// TIA Portal project "ESTHER_Gas_v4.0_4" (V13) (continued)
       #DATA_ADDR := "MB_AD_COUNTER_RST_ENABL";
       #DATA_INT_PTR.DATA[0] := "MB_VAL_COUNT_RST_ENABL";
   END_IF;
   IF #"STEP" = 44 THEN
       #DATA_ADDR := "MB_AD_COUNTER_UNIT_IDX";
       #DATA_INT_PTR.DATA[0] := 0;   // Unit: ln
   END_IF;
   IF #"STEP" = 45 THEN
       #DATA_ADDR := "MB_AD_COUNTER_SP_MODE";
       #DATA_INT_PTR.DATA[0] := "MB_VAL_COUNT_SP_MODE_CHANGE";
   END_IF;
   IF #"STEP" = 46 THEN
       #DATA_ADDR := "MB_AD_COUNTER_NEW_SP";
       #DATA_INT_PTR.DATA[0] := 0;
   END_IF;
   IF #"STEP" = 47 THEN
       #DATA_ADDR := "MB_AD_RESET";
       #DATA_INT_PTR.DATA[0] := 0;
   END_IF;
   IF #"STEP" = 48 THEN
       #DATA_ADDR := "MB_AD_RESET";
       #DATA_INT_PTR.DATA[0] := 3;
   END_IF;
   IF #"STEP" = 49 THEN
       #DATA_ADDR := "MB_AD_COUNTER_MODE";
       #DATA_INT_PTR.DATA[0] := "MB_VAL_COUNT_MODE_UP_LIMIT";
   END_IF;
   IF #"STEP" = 50 THEN
       #MB_MODE := 1;
       #DATA_LEN := 1;
       #DATA_ADDR := #MB_AD_CONTROL_MODE;
       #DATA_INT_PTR.DATA[0] := #MFC_MODE_SP;   // SET ControlMode
   END_IF;
   IF #"STEP" = 60 THEN
       #MB_MODE := 1;
       #DATA_LEN := 1;
       #DATA_ADDR := #MB_AD_CONTROL_MODE;
       #DATA_INT_PTR.DATA[0] := 0;   // SET ControlMode Bus
   END_IF;
   IF #"STEP" = 63 THEN
       #MB_MODE := 1;
       #DATA_LEN := 1;
       #DATA_ADDR := #MB_AD_CONTROL_MODE;
       #DATA_INT_PTR.DATA[0] := 3;   // SET ControlMode Close
   END_IF;
   IF #"STEP" = 68 THEN
       #MB_MODE := 1;
       #DATA_LEN := 1;
       #DATA_ADDR := #MB_AD_CONTROL_MODE;
       #DATA_INT_PTR.DATA[0] := 8;   // SET ControlMode Open
   END_IF;
   IF #"STEP" = 80 THEN
       #MB_MODE := 1;
       #DATA_LEN := 1;
       #DATA_ADDR := "MB_AD_SETPOINT";
       #DATA_INT_PTR.DATA[0] := #MFC_Setpoint;   // Set Setpoint
   END_IF;
END_REGION
END_FUNCTION_BLOCK

FUNCTION_BLOCK "ETAPA_1_HE_NOK"   // FB3, LAD
{ S7_Optimized_Access := 'FALSE' }
VERSION : 0.1
// Inertização da Câmara de testes com Helio.
BEGIN

REGION Network 1
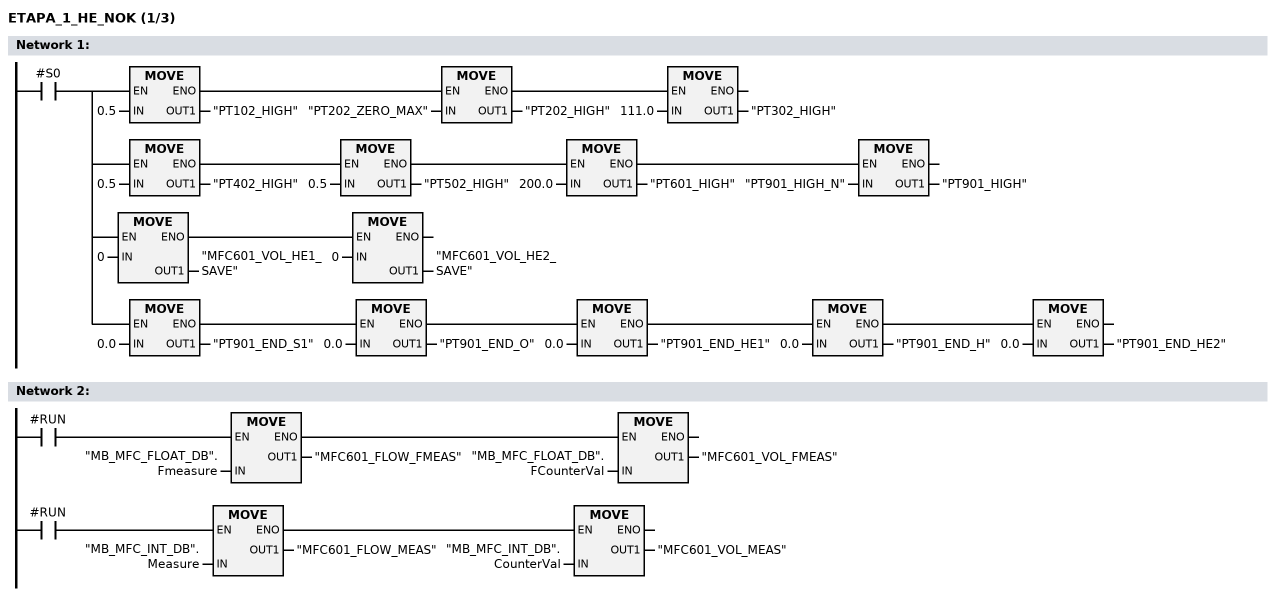
   RUNG wire#powerrail
      Contact( #S0 )
      wire#w1
      { S7_GenerateENO := "TRUE" } Move(in := 0.5, out1 => "PT102_HIGH")
      { S7_GenerateENO := "TRUE" } Move(in := "PT202_ZERO_MAX", out1 => "PT202_HIGH")
      { S7_GenerateENO := "TRUE" } Move(in := 111.0, out1 => "PT302_HIGH")
   END_RUNG
   RUNG wire#w1
      { S7_GenerateENO := "TRUE" } Move(in := 0.5, out1 => "PT402_HIGH")
      { S7_GenerateENO := "TRUE" } Move(in := 0.5, out1 => "PT502_HIGH")
      { S7_GenerateENO := "TRUE" } Move(in := 200.0, out1 => "PT601_HIGH")
      { S7_GenerateENO := "TRUE" } Move(in := "PT901_HIGH_N", out1 => "PT901_HIGH")
   END_RUNG
   RUNG wire#w1
      { S7_GenerateENO := "TRUE" } Move(in := 0, out1 => "MFC601_VOL_HE1_SAVE")
      { S7_GenerateENO := "TRUE" } Move(in := 0, out1 => "MFC601_VOL_HE2_SAVE")
   END_RUNG
   RUNG wire#w1
      { S7_GenerateENO := "TRUE" } Move(in := 0.0, out1 => "PT901_END_S1")
      { S7_GenerateENO := "TRUE" } Move(in := 0.0, out1 => "PT901_END_O")
      { S7_GenerateENO := "TRUE" } Move(in := 0.0, out1 => "PT901_END_HE1")
      { S7_GenerateENO := "TRUE" } Move(in := 0.0, out1 => "PT901_END_H")
      { S7_GenerateENO := "TRUE" } Move(in := 0.0, out1 => "PT901_END_HE2")
   END_RUNG
   // the same network as SCL:
   // ENO of a box is taken as its EN; it also drops when the box reports an error
   IF #S0 THEN
       "PT102_HIGH" := 0.5;
       "PT202_HIGH" := "PT202_ZERO_MAX";
       "PT302_HIGH" := 111.0;
       "PT402_HIGH" := 0.5;
       "PT502_HIGH" := 0.5;
       "PT601_HIGH" := 200.0;
       "PT901_HIGH" := "PT901_HIGH_N";
       "MFC601_VOL_HE1_SAVE" := 0;
       "MFC601_VOL_HE2_SAVE" := 0;
       "PT901_END_S1" := 0.0;
       "PT901_END_O" := 0.0;
       "PT901_END_HE1" := 0.0;
       "PT901_END_H" := 0.0;
       "PT901_END_HE2" := 0.0;
   END_IF;
END_REGION

REGION Network 2
   RUNG wire#powerrail
      Contact( #RUN )
      { S7_GenerateENO := "TRUE" } Move(in := "MB_MFC_FLOAT_DB".Fmeasure, out1 => "MFC601_FLOW_FMEAS")
      { S7_GenerateENO := "TRUE" } Move(in := "MB_MFC_FLOAT_DB".FCounterVal, out1 => "MFC601_VOL_FMEAS")
   END_RUNG
   RUNG wire#powerrail
      Contact( #RUN )
      { S7_GenerateENO := "TRUE" } Move(in := "MB_MFC_INT_DB".Measure, out1 => "MFC601_FLOW_MEAS")
      { S7_GenerateENO := "TRUE" } Move(in := "MB_MFC_INT_DB".CounterVal, out1 => "MFC601_VOL_MEAS")
   END_RUNG
   // the same network as SCL:
   // ENO of a box is taken as its EN; it also drops when the box reports an error
   IF #RUN THEN
       "MFC601_FLOW_FMEAS" := "MB_MFC_FLOAT_DB".Fmeasure;
       "MFC601_VOL_FMEAS" := "MB_MFC_FLOAT_DB".FCounterVal;
       "MFC601_FLOW_MEAS" := "MB_MFC_INT_DB".Measure;
       "MFC601_VOL_MEAS" := "MB_MFC_INT_DB".CounterVal;
   END_IF;
END_REGION

REGION Network 3
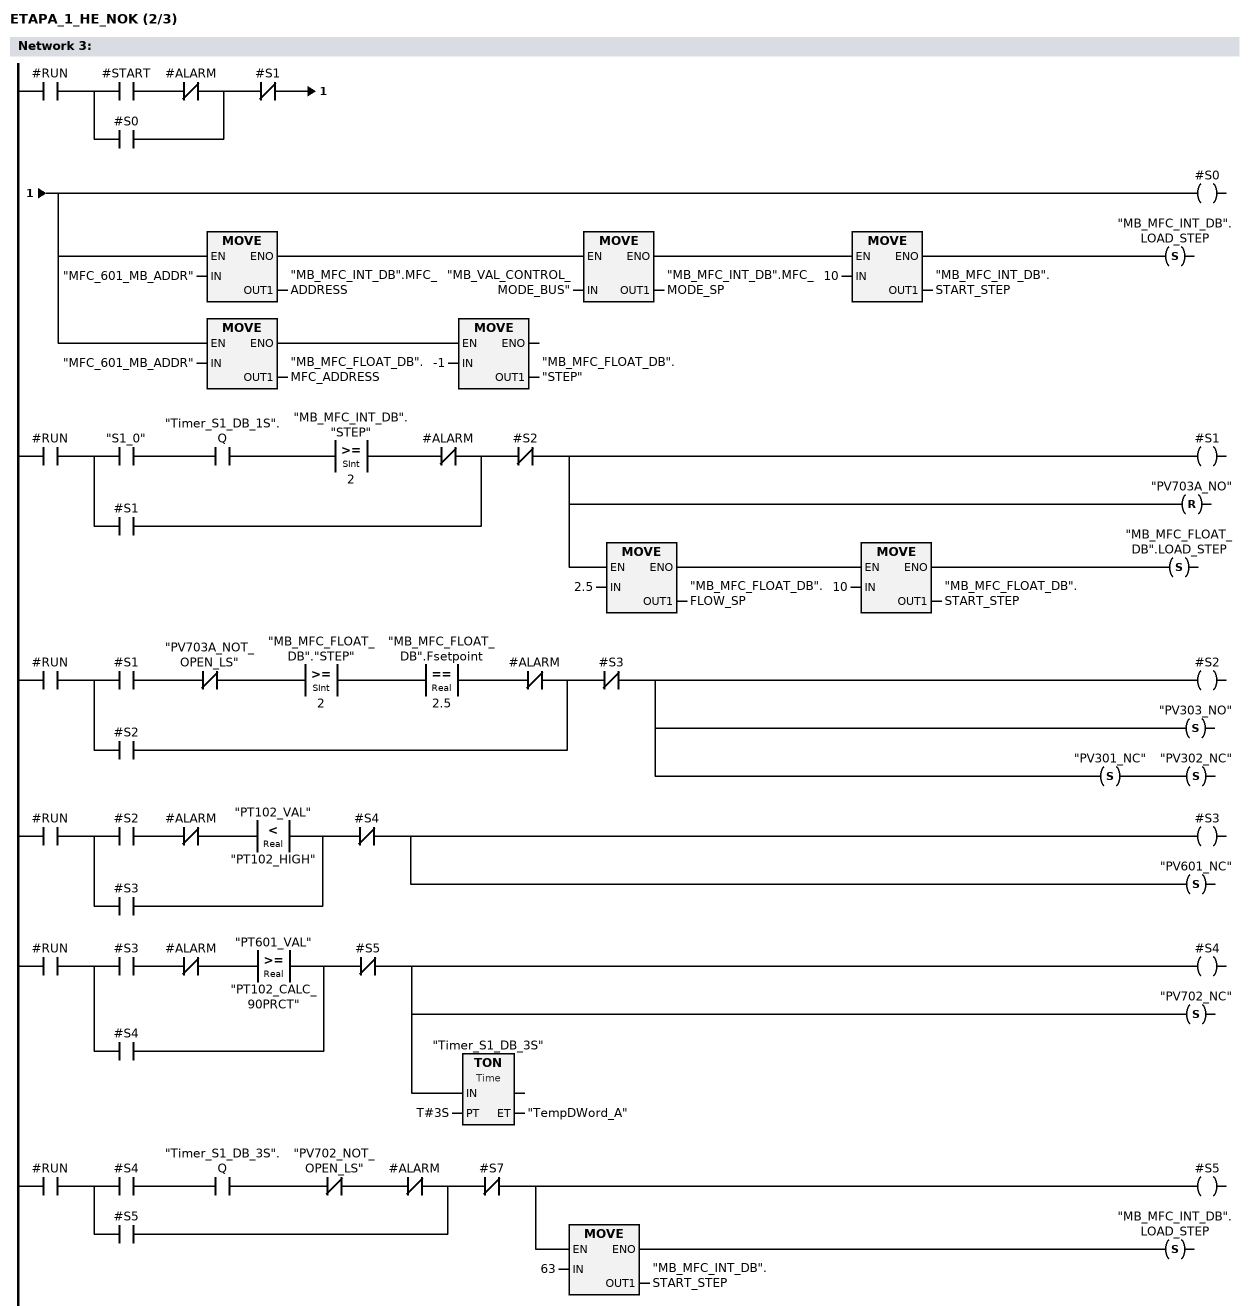
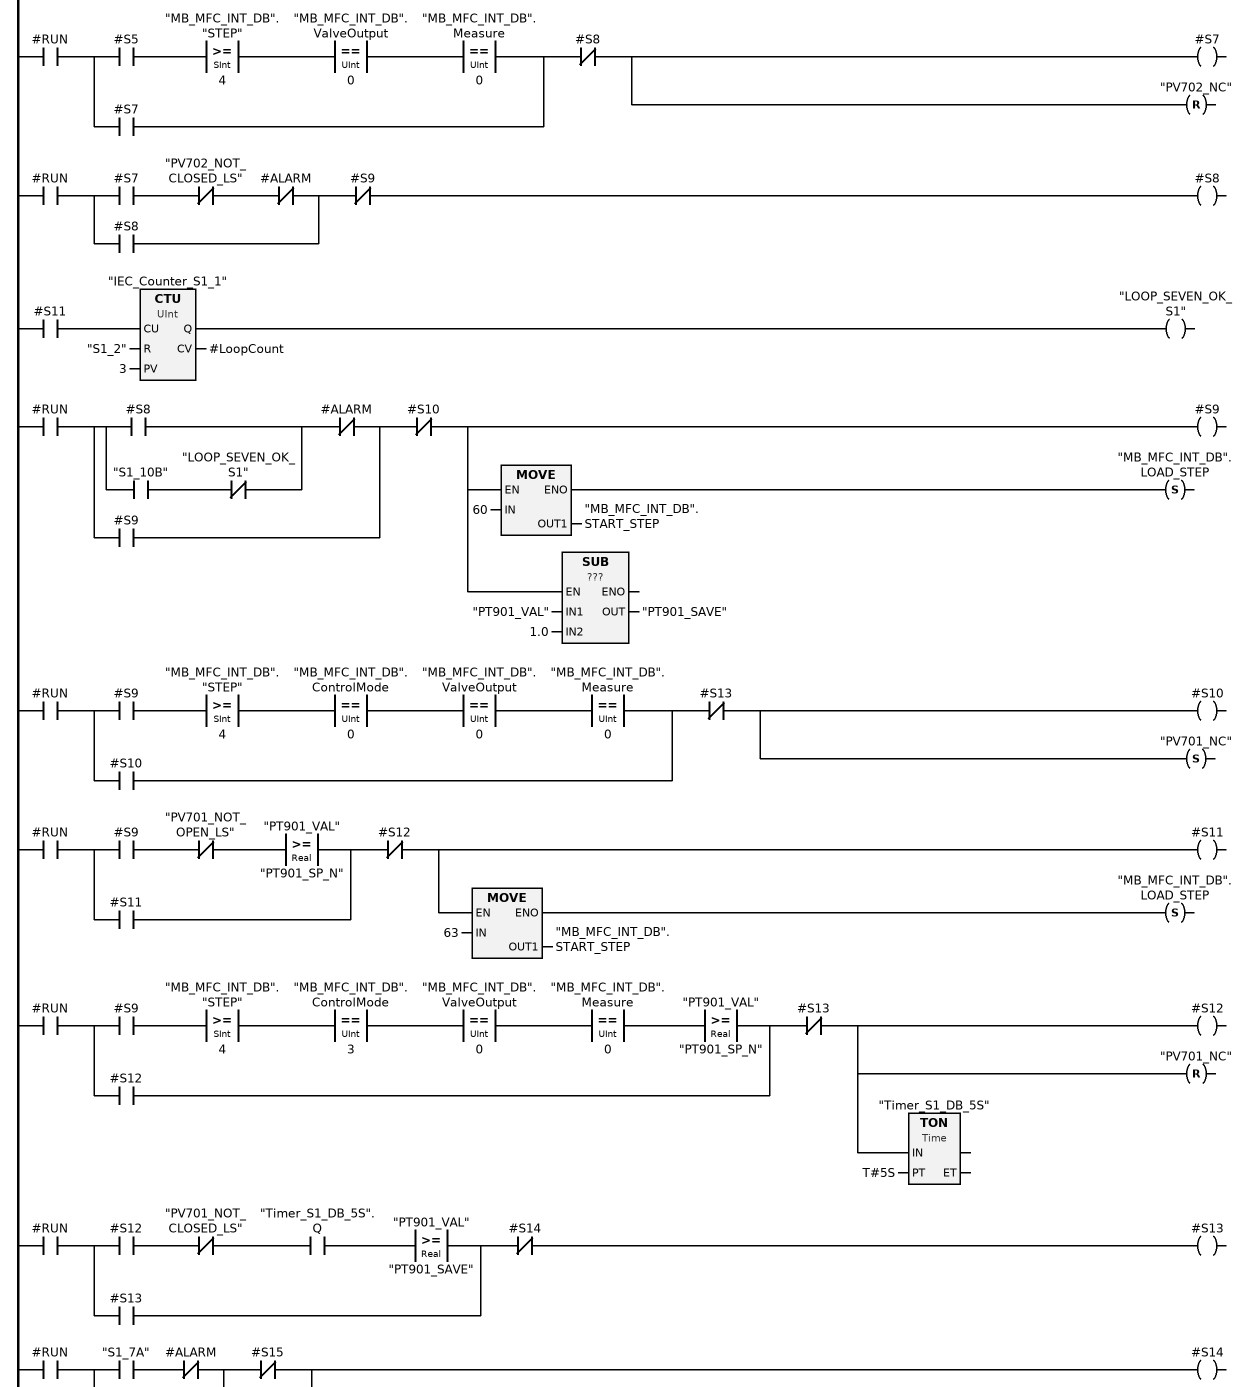
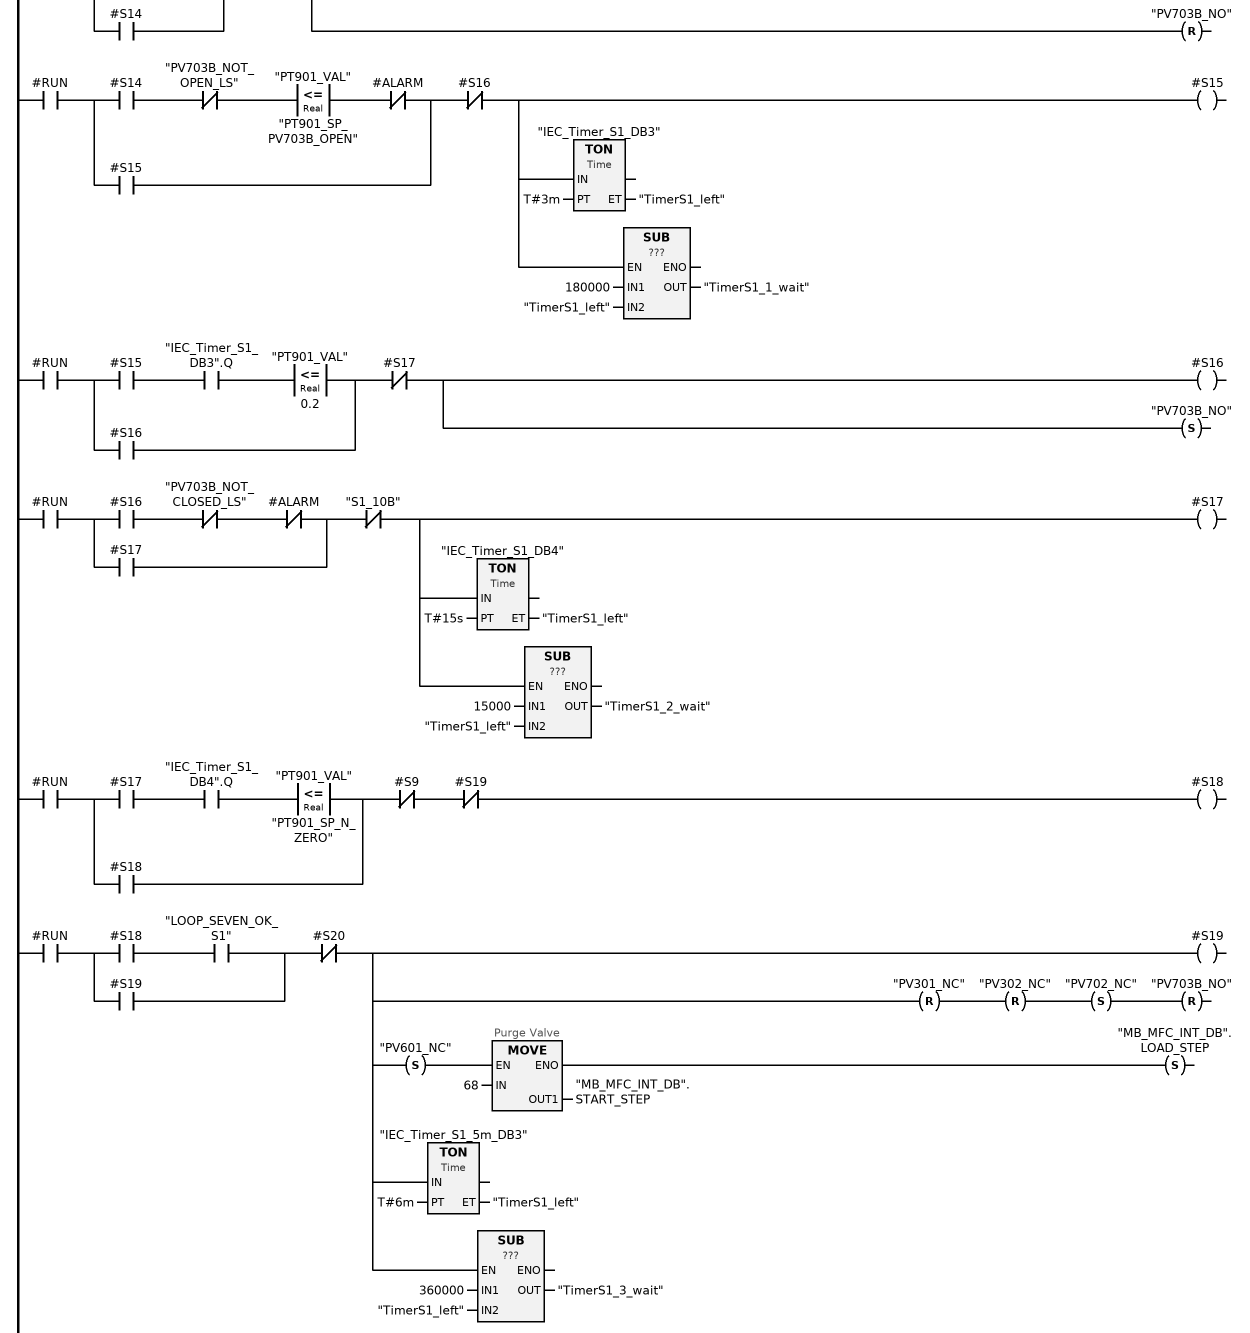
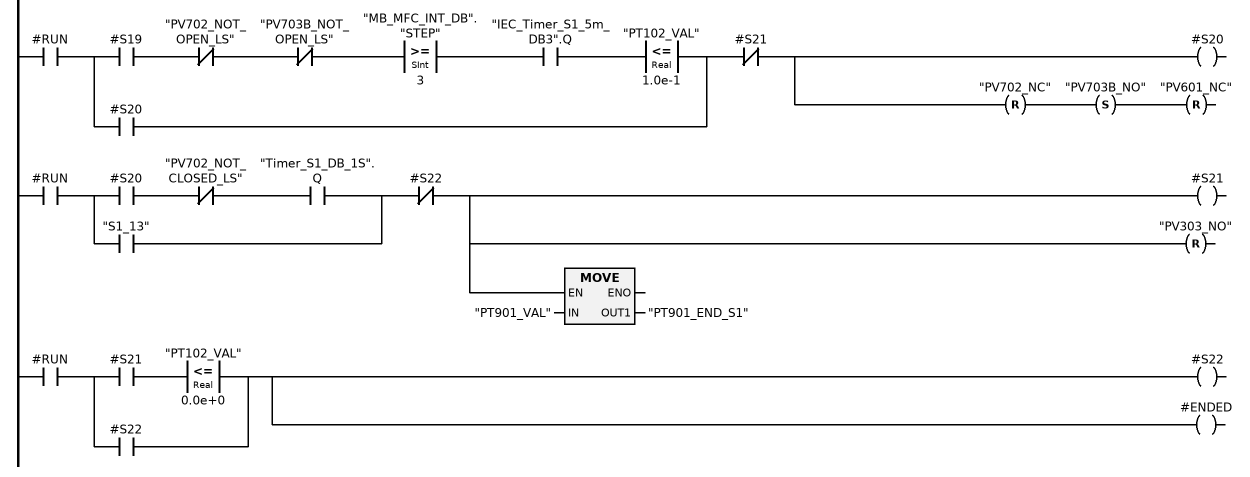
   #S0 := #RUN AND ((#START AND NOT #ALARM) OR #S0) AND NOT #S1;
   IF #S0 THEN
       "MB_MFC_INT_DB".MFC_ADDRESS := "MFC_601_MB_ADDR";
       "MB_MFC_INT_DB".MFC_MODE_SP := "MB_VAL_CONTROL_MODE_BUS";
       "MB_MFC_INT_DB".START_STEP := 10;
       "MB_MFC_INT_DB".LOAD_STEP := TRUE;
       "MB_MFC_FLOAT_DB".MFC_ADDRESS := "MFC_601_MB_ADDR";
       "MB_MFC_FLOAT_DB"."STEP" := -1;
   END_IF;
   #S1 := #RUN AND (("S1_0" AND "Timer_S1_DB_1S".Q AND ("MB_MFC_INT_DB"."STEP" >= 2) AND NOT #ALARM) OR #S1) AND NOT #S2;
   IF #S1 THEN
       "PV703A_NO" := FALSE;
       "MB_MFC_FLOAT_DB".FLOW_SP := 2.5;
       "MB_MFC_FLOAT_DB".START_STEP := 10;
       "MB_MFC_FLOAT_DB".LOAD_STEP := TRUE;
   END_IF;
   #S2 := #RUN AND ((#S1 AND NOT "PV703A_NOT_OPEN_LS" AND ("MB_MFC_FLOAT_DB"."STEP" >= 2) AND ("MB_MFC_FLOAT_DB".Fsetpoint = 2.5) AND NOT #ALARM) OR #S2) AND NOT #S3;
   IF #S2 THEN
       "PV303_NO" := TRUE;
       "PV301_NC" := TRUE;
       "PV302_NC" := TRUE;
   END_IF;
   #S3 := #RUN AND ((#S2 AND NOT #ALARM AND ("PT102_VAL" < "PT102_HIGH")) OR #S3) AND NOT #S4;
   IF #S3 THEN "PV601_NC" := TRUE; END_IF;
   #S4 := #RUN AND ((#S3 AND NOT #ALARM AND ("PT601_VAL" >= "PT102_CALC_90PRCT")) OR #S4) AND NOT #S5;
   IF #S4 THEN "PV702_NC" := TRUE; END_IF;
   "Timer_S1_DB_3S".TON(IN := #S4, PT := T#3S, ET => "TempDWord_A");
   #S5 := #RUN AND ((#S4 AND "Timer_S1_DB_3S".Q AND NOT "PV702_NOT_OPEN_LS" AND NOT #ALARM) OR #S5) AND NOT #S7;
   IF #S5 THEN
       "MB_MFC_INT_DB".START_STEP := 63;
       "MB_MFC_INT_DB".LOAD_STEP := TRUE;
   END_IF;
   #S7 := #RUN AND ((#S5 AND ("MB_MFC_INT_DB"."STEP" >= 4) AND ("MB_MFC_INT_DB".ValveOutput = 0) AND ("MB_MFC_INT_DB".Measure = 0)) OR #S7) AND NOT #S8;
   IF #S7 THEN "PV702_NC" := FALSE; END_IF;
   #S8 := #RUN AND ((#S7 AND NOT "PV702_NOT_CLOSED_LS" AND NOT #ALARM) OR #S8) AND NOT #S9;
   "IEC_Counter_S1_1".CTU(CU := #S11, R := "S1_2", PV := 3, CV => #LoopCount);
   "LOOP_SEVEN_OK_S1" := "IEC_Counter_S1_1".Q;
   #S9 := #RUN AND (((#S8 OR ("S1_10B" AND NOT "LOOP_SEVEN_OK_S1")) AND NOT #ALARM) OR #S9) AND NOT #S10;
   IF #S9 THEN
       "MB_MFC_INT_DB".START_STEP := 60;
       "MB_MFC_INT_DB".LOAD_STEP := TRUE;
       "PT901_SAVE" := "PT901_VAL" - 1.0;
   END_IF;
   #S10 := #RUN AND ((#S9 AND ("MB_MFC_INT_DB"."STEP" >= 4) AND ("MB_MFC_INT_DB".ControlMode = 0) AND ("MB_MFC_INT_DB".ValveOutput = 0) AND ("MB_MFC_INT_DB".Measure = 0)) OR #S10) AND NOT #S13;
   IF #S10 THEN "PV701_NC" := TRUE; END_IF;
   #S11 := #RUN AND ((#S9 AND NOT "PV701_NOT_OPEN_LS" AND ("PT901_VAL" >= "PT901_SP_N")) OR #S11) AND NOT #S12;
   IF #S11 THEN
       "MB_MFC_INT_DB".START_STEP := 63;
       "MB_MFC_INT_DB".LOAD_STEP := TRUE;
   END_IF;
   #S12 := #RUN AND ((#S9 AND ("MB_MFC_INT_DB"."STEP" >= 4) AND ("MB_MFC_INT_DB".ControlMode = 3) AND ("MB_MFC_INT_DB".ValveOutput = 0) AND ("MB_MFC_INT_DB".Measure = 0) AND ("PT901_VAL" >= "PT901_SP_N")) OR #S12) AND NOT #S13;
   IF #S12 THEN "PV701_NC" := FALSE; END_IF;
   "Timer_S1_DB_5S".TON(IN := #S12, PT := T#5S);
   #S13 := #RUN AND ((#S12 AND NOT "PV701_NOT_CLOSED_LS" AND "Timer_S1_DB_5S".Q AND ("PT901_VAL" >= "PT901_SAVE")) OR #S13) AND NOT #S14;
   #S14 := #RUN AND (("S1_7A" AND NOT #ALARM) OR #S14) AND NOT #S15;
   IF #S14 THEN "PV703B_NO" := FALSE; END_IF;
   #S15 := #RUN AND ((#S14 AND NOT "PV703B_NOT_OPEN_LS" AND ("PT901_VAL" <= "PT901_SP_PV703B_OPEN") AND NOT #ALARM) OR #S15) AND NOT #S16;
   "IEC_Timer_S1_DB3".TON(IN := #S15, PT := T#3m, ET => "TimerS1_left");
   IF #S15 THEN "TimerS1_1_wait" := 180000 - "TimerS1_left"; END_IF;
   #S16 := #RUN AND ((#S15 AND "IEC_Timer_S1_DB3".Q AND ("PT901_VAL" <= 0.2)) OR #S16) AND NOT #S17;
   IF #S16 THEN "PV703B_NO" := TRUE; END_IF;
   #S17 := #RUN AND ((#S16 AND NOT "PV703B_NOT_CLOSED_LS" AND NOT #ALARM) OR #S17) AND NOT "S1_10B";
   "IEC_Timer_S1_DB4".TON(IN := #S17, PT := T#15s, ET => "TimerS1_left");
   IF #S17 THEN "TimerS1_2_wait" := 15000 - "TimerS1_left"; END_IF;
   #S18 := #RUN AND ((#S17 AND "IEC_Timer_S1_DB4".Q AND ("PT901_VAL" <= "PT901_SP_N_ZERO")) OR #S18) AND NOT #S9 AND NOT #S19;
   #S19 := #RUN AND ((#S18 AND "LOOP_SEVEN_OK_S1") OR #S19) AND NOT #S20;
   IF #S19 THEN
       "PV301_NC" := FALSE;
       "PV302_NC" := FALSE;
       "PV702_NC" := TRUE;
       "PV703B_NO" := FALSE;
       "PV601_NC" := TRUE;
       "MB_MFC_INT_DB".START_STEP := 68;   // Purge Valve
       "MB_MFC_INT_DB".LOAD_STEP := TRUE;
   END_IF;
   "IEC_Timer_S1_5m_DB3".TON(IN := #S19, PT := T#6m, ET => "TimerS1_left");
   IF #S19 THEN "TimerS1_3_wait" := 360000 - "TimerS1_left"; END_IF;
   #S20 := #RUN AND ((#S19 AND NOT "PV702_NOT_OPEN_LS" AND NOT "PV703B_NOT_OPEN_LS" AND ("MB_MFC_INT_DB"."STEP" >= 3) AND "IEC_Timer_S1_5m_DB3".Q AND ("PT102_VAL" <= 1.0e-1)) OR #S20) AND NOT #S21;
   IF #S20 THEN
       "PV702_NC" := FALSE;
       "PV703B_NO" := TRUE;
       "PV601_NC" := FALSE;
   END_IF;
   #S21 := #RUN AND ((#S20 AND NOT "PV702_NOT_CLOSED_LS" AND "Timer_S1_DB_1S".Q) OR "S1_13") AND NOT #S22;
   IF #S21 THEN
       "PV303_NO" := FALSE;
       "PT901_END_S1" := "PT901_VAL";
   END_IF;
   #S22 := #RUN AND ((#S21 AND ("PT102_VAL" <= 0.0e+0)) OR #S22);
   #ENDED := #S22;
END_REGION

REGION Network 4
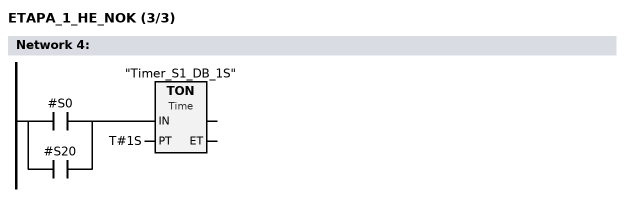
   "Timer_S1_DB_1S".TON(IN := #S0 OR #S20, PT := T#1S);
END_REGION
END_FUNCTION_BLOCK

FUNCTION "ETAPA_1_N" : Void   // FC1, LAD
{ S7_Optimized_Access := 'FALSE' }
VERSION : 0.1
// Inertização da Câmara de testes com N2. Max SP N2 =2.5 Bar. Loop times = 2 (testing)
// S!_10 A ->10s
BEGIN

REGION Network 1: Alarm Set points
   // Alarm Set points of this step
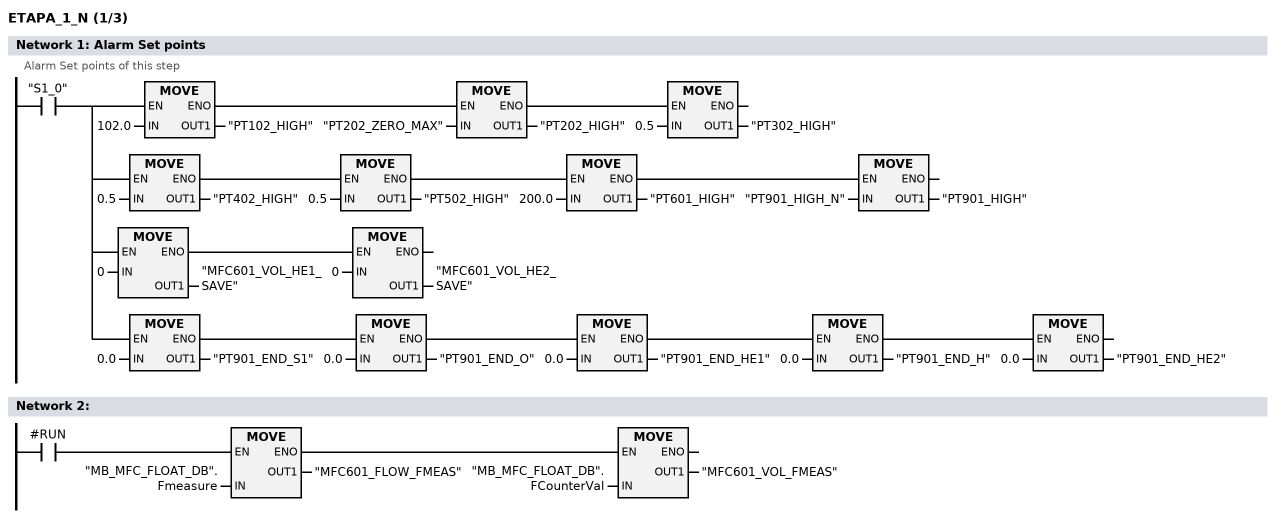
   RUNG wire#powerrail
      Contact( "S1_0" )
      wire#w1
      { S7_GenerateENO := "TRUE" } Move(in := 102.0, out1 => "PT102_HIGH")
      { S7_GenerateENO := "TRUE" } Move(in := "PT202_ZERO_MAX", out1 => "PT202_HIGH")
      { S7_GenerateENO := "TRUE" } Move(in := 0.5, out1 => "PT302_HIGH")
   END_RUNG
   RUNG wire#w1
      { S7_GenerateENO := "TRUE" } Move(in := 0.5, out1 => "PT402_HIGH")
      { S7_GenerateENO := "TRUE" } Move(in := 0.5, out1 => "PT502_HIGH")
      { S7_GenerateENO := "TRUE" } Move(in := 200.0, out1 => "PT601_HIGH")
      { S7_GenerateENO := "TRUE" } Move(in := "PT901_HIGH_N", out1 => "PT901_HIGH")
   END_RUNG
   RUNG wire#w1
      { S7_GenerateENO := "TRUE" } Move(in := 0, out1 => "MFC601_VOL_HE1_SAVE")
      { S7_GenerateENO := "TRUE" } Move(in := 0, out1 => "MFC601_VOL_HE2_SAVE")
   END_RUNG
   RUNG wire#w1
      { S7_GenerateENO := "TRUE" } Move(in := 0.0, out1 => "PT901_END_S1")
      { S7_GenerateENO := "TRUE" } Move(in := 0.0, out1 => "PT901_END_O")
      { S7_GenerateENO := "TRUE" } Move(in := 0.0, out1 => "PT901_END_HE1")
      { S7_GenerateENO := "TRUE" } Move(in := 0.0, out1 => "PT901_END_H")
      { S7_GenerateENO := "TRUE" } Move(in := 0.0, out1 => "PT901_END_HE2")
   END_RUNG
   // the same network as SCL:
   // ENO of a box is taken as its EN; it also drops when the box reports an error
   IF "S1_0" THEN
       "PT102_HIGH" := 102.0;
       "PT202_HIGH" := "PT202_ZERO_MAX";
       "PT302_HIGH" := 0.5;
       "PT402_HIGH" := 0.5;
       "PT502_HIGH" := 0.5;
       "PT601_HIGH" := 200.0;
       "PT901_HIGH" := "PT901_HIGH_N";
       "MFC601_VOL_HE1_SAVE" := 0;
       "MFC601_VOL_HE2_SAVE" := 0;
       "PT901_END_S1" := 0.0;
       "PT901_END_O" := 0.0;
       "PT901_END_HE1" := 0.0;
       "PT901_END_H" := 0.0;
       "PT901_END_HE2" := 0.0;
   END_IF;
END_REGION

REGION Network 2
   RUNG wire#powerrail
      Contact( #RUN )
      { S7_GenerateENO := "TRUE" } Move(in := "MB_MFC_FLOAT_DB".Fmeasure, out1 => "MFC601_FLOW_FMEAS")
      { S7_GenerateENO := "TRUE" } Move(in := "MB_MFC_FLOAT_DB".FCounterVal, out1 => "MFC601_VOL_FMEAS")
   END_RUNG
   // the same network as SCL:
   // ENO of a box is taken as its EN; it also drops when the box reports an error
   IF #RUN THEN
       "MFC601_FLOW_FMEAS" := "MB_MFC_FLOAT_DB".Fmeasure;
       "MFC601_VOL_FMEAS" := "MB_MFC_FLOAT_DB".FCounterVal;
   END_IF;
END_REGION

REGION Network 3